   2383: 'Carrier 37 Encoder Comm Fault', class No Acknowledgement, trigger "DB302_HMI_Faults_Carrier37_Faults_0" bit 14
   2384: 'Carrier 37 HMI Comm Fault', class No Acknowledgement, trigger "DB302_HMI_Faults_Carrier37_Faults_0" bit 15
   2385: 'Carrier 37 Crash Detection Fault', class No Acknowledgement, trigger "DB302_HMI_Faults_Carrier37_Faults_1" bit 0
   2386: 'Carrier 37 Carrier Number Invalid', class No Acknowledgement, trigger "DB302_HMI_Faults_Carrier37_Faults_1" bit 1
   2387: 'Carrier 37 Drive: PROFINET configuration error', class No Acknowledgement, trigger "DB302_HMI_Faults_Carrier37_Faults_1" bit 2
   2388: 'Carrier 37 Drive: Error internal communications', class No Acknowledgement, trigger "DB302_HMI_Faults_Carrier37_Faults_1" bit 3
   2389: 'Carrier 37 Drive: Motor overtemperature', class No Acknowledgement, trigger "DB302_HMI_Faults_Carrier37_Faults_1" bit 4
   2390: 'Carrier 37 Drive: Motor overcurrent', class No Acknowledgement, trigger "DB302_HMI_Faults_Carrier37_Faults_1" bit 5
   2391: 'Carrier 37 Drive: Infeed or power unit not ready', class No Acknowledgement, trigger "DB302_HMI_Faults_Carrier37_Faults_1" bit 6
   2392: 'Carrier 37 Drive: Short-circuit/ground fault detected', class No Acknowledgement, trigger "DB302_HMI_Faults_Carrier37_Faults_1" bit 7
   2393: 'Carrier 37 Drive: PROFINET Setpoint timeout', class No Acknowledgement, trigger "DB302_HMI_Faults_Carrier37_Faults_1" bit 8
   2394: 'Carrier 37 Power unit: Overcurrent', class No Acknowledgement, trigger "DB302_HMI_Faults_Carrier37_Faults_1" bit 9
   2395: 'Carrier 37 Power unit: DC link voltage overvoltage', class No Acknowledgement, trigger "DB302_HMI_Faults_Carrier37_Faults_1" bit 10
   2396: 'Carrier 37 Power unit: DC link voltage undervoltage', class No Acknowledgement, trigger "DB302_HMI_Faults_Carrier37_Faults_1" bit 11
   2397: 'Carrier 37 Power unit: Line phase failure in main circuit', class No Acknowledgement, trigger "DB302_HMI_Faults_Carrier37_Faults_1" bit 12
   2398: 'Carrier 37 Power unit: Phase failure motor cable', class No Acknowledgement, trigger "DB302_HMI_Faults_Carrier37_Faults_1" bit 13
   2399: 'Carrier 37 Power unit: Ground fault', class No Acknowledgement, trigger "DB302_HMI_Faults_Carrier37_Faults_1" bit 14
   2400: 'Spare_Fault_2400', class No Acknowledgement, trigger "DB302_HMI_Faults_Carrier37_Faults_1" bit 15
   2401: 'Carrier 37 Motion Off Fault', class No Acknowledgement, trigger "DB302_HMI_Faults_Carrier37_Faults_2" bit 0
   2402: 'Carrier 37 Motion On Fault', class No Acknowledgement, trigger "DB302_HMI_Faults_Carrier37_Faults_2" bit 1
   2403: 'Carrier 37 Spacing Fault', class No Acknowledgement, trigger "DB302_HMI_Faults_Carrier37_Faults_2" bit 2
   2404: 'Carrier 37 Duplicate Carrier Number Fault', class No Acknowledgement, trigger "DB302_HMI_Faults_Carrier37_Faults_2" bit 3
   2405: 'Spare_Fault_2405', class No Acknowledgement, trigger "DB302_HMI_Faults_Carrier37_Faults_2" bit 4
   2406: 'Spare_Fault_2406', class No Acknowledgement, trigger "DB302_HMI_Faults_Carrier37_Faults_2" bit 5
   2407: 'Spare_Fault_2407', class No Acknowledgement, trigger "DB302_HMI_Faults_Carrier37_Faults_2" bit 6
   2408: 'Spare_Fault_2408', class No Acknowledgement, trigger "DB302_HMI_Faults_Carrier37_Faults_2" bit 7
   2409: 'Spare_Fault_2409', class No Acknowledgement, trigger "DB302_HMI_Faults_Carrier37_Faults_2" bit 8
   2410: 'Spare_Fault_2410', class No Acknowledgement, trigger "DB302_HMI_Faults_Carrier37_Faults_2" bit 9
   2411: 'Spare_Fault_2411', class No Acknowledgement, trigger "DB302_HMI_Faults_Carrier37_Faults_2" bit 10
   2412: 'Spare_Fault_2412', class No Acknowledgement, trigger "DB302_HMI_Faults_Carrier37_Faults_2" bit 11
   2413: 'Spare_Fault_2413', class No Acknowledgement, trigger "DB302_HMI_Faults_Carrier37_Faults_2" bit 12
   2414: 'Spare_Fault_2414', class No Acknowledgement, trigger "DB302_HMI_Faults_Carrier37_Faults_2" bit 13
   2415: 'Spare_Fault_2415', class No Acknowledgement, trigger "DB302_HMI_Faults_Carrier37_Faults_2" bit 14
   2416: 'Spare_Fault_2416', class No Acknowledgement, trigger "DB302_HMI_Faults_Carrier37_Faults_2" bit 15
   2417: 'Spare_Fault_2417', class No Acknowledgement, trigger "DB302_HMI_Faults_Carrier37_Faults_3" bit 0
   2418: 'Spare_Fault_2418', class No Acknowledgement, trigger "DB302_HMI_Faults_Carrier37_Faults_3" bit 1
   2419: 'Spare_Fault_2419', class No Acknowledgement, trigger "DB302_HMI_Faults_Carrier37_Faults_3" bit 2
   2420: 'Spare_Fault_2420', class No Acknowledgement, trigger "DB302_HMI_Faults_Carrier37_Faults_3" bit 3
   2421: 'Spare_Fault_2421', class No Acknowledgement, trigger "DB302_HMI_Faults_Carrier37_Faults_3" bit 4
   2422: 'Spare_Fault_2422', class No Acknowledgement, trigger "DB302_HMI_Faults_Carrier37_Faults_3" bit 5
   2423: 'Spare_Fault_2423', class No Acknowledgement, trigger "DB302_HMI_Faults_Carrier37_Faults_3" bit 6
   2424: 'Spare_Fault_2424', class No Acknowledgement, trigger "DB302_HMI_Faults_Carrier37_Faults_3" bit 7
   2425: 'Spare_Fault_2425', class No Acknowledgement, trigger "DB302_HMI_Faults_Carrier37_Faults_3" bit 8
   2426: 'Spare_Fault_2426', class No Acknowledgement, trigger "DB302_HMI_Faults_Carrier37_Faults_3" bit 9
   2427: 'Spare_Fault_2427', class No Acknowledgement, trigger "DB302_HMI_Faults_Carrier37_Faults_3" bit 10
   2428: 'Spare_Fault_2428', class No Acknowledgement, trigger "DB302_HMI_Faults_Carrier37_Faults_3" bit 11
   2429: 'Spare_Fault_2429', class No Acknowledgement, trigger "DB302_HMI_Faults_Carrier37_Faults_3" bit 12
   2430: 'Spare_Fault_2430', class No Acknowledgement, trigger "DB302_HMI_Faults_Carrier37_Faults_3" bit 13
   2431: 'Spare_Fault_2431', class No Acknowledgement, trigger "DB302_HMI_Faults_Carrier37_Faults_3" bit 14
   2432: 'Spare_Fault_2432', class No Acknowledgement, trigger "DB302_HMI_Faults_Carrier37_Faults_3" bit 15
   2433: 'Carrier 38 Disconnect Open Power Fault DI11.0', class No Acknowledgement, trigger "DB302_HMI_Faults_Carrier38_Faults_0" bit 0
   2434: 'Carrier 38 Drive Profinet Comm Fault', class No Acknowledgement, trigger "DB302_HMI_Faults_Carrier38_Faults_0" bit 1
   2435: 'Carrier 38 Production Stop Not Reset', class No Acknowledgement, trigger "DB302_HMI_Faults_Carrier38_Faults_0" bit 2
   2436: 'Carrier 38 CB02122 Tripped', class No Acknowledgement, trigger "DB302_HMI_Faults_Carrier38_Faults_0" bit 3
   2437: 'Carrier 38 CB02123 Tripped', class No Acknowledgement, trigger "DB302_HMI_Faults_Carrier38_Faults_0" bit 4
   2438: 'Carrier 38 AUX1 CB Tripped', class No Acknowledgement, trigger "DB302_HMI_Faults_Carrier38_Faults_0" bit 5
   2439: 'Carrier 38 AUX2 CB Tripped', class No Acknowledgement, trigger "DB302_HMI_Faults_Carrier38_Faults_0" bit 6
   2440: 'Carrier 38 PLC Not Communicating', class No Acknowledgement, trigger "DB302_HMI_Faults_Carrier38_Faults_0" bit 7
   2441: 'Carrier 38 Safe Input Card Fault', class No Acknowledgement, trigger "DB302_HMI_Faults_Carrier38_Faults_0" bit 8
   2442: 'Carrier 38 Safe Output Card Fault', class No Acknowledgement, trigger "DB302_HMI_Faults_Carrier38_Faults_0" bit 9
   2443: 'Carrier 38 Standard Input Card Fault', class No Acknowledgement, trigger "DB302_HMI_Faults_Carrier38_Faults_0" bit 10
   2444: 'Carrier 38 Standard Output Card Fault', class No Acknowledgement, trigger "DB302_HMI_Faults_Carrier38_Faults_0" bit 11
   2445: 'Carrier 38 Encoder Position Fault', class No Acknowledgement, trigger "DB302_HMI_Faults_Carrier38_Faults_0" bit 12
   2446: 'Carrier 38 Encoder Internal Error', class No Acknowledgement, trigger "DB302_HMI_Faults_Carrier38_Faults_0" bit 13
   2447: 'Carrier 38 Encoder Comm Fault', class No Acknowledgement, trigger "DB302_HMI_Faults_Carrier38_Faults_0" bit 14
   2448: 'Carrier 38 HMI Comm Fault', class No Acknowledgement, trigger "DB302_HMI_Faults_Carrier38_Faults_0" bit 15
   2449: 'Carrier 38 Crash Detection Fault', class No Acknowledgement, trigger "DB302_HMI_Faults_Carrier38_Faults_1" bit 0
   2450: 'Carrier 38 Carrier Number Invalid', class No Acknowledgement, trigger "DB302_HMI_Faults_Carrier38_Faults_1" bit 1
   2451: 'Carrier 38 Drive: PROFINET configuration error', class No Acknowledgement, trigger "DB302_HMI_Faults_Carrier38_Faults_1" bit 2
   2452: 'Carrier 38 Drive: Error internal communications', class No Acknowledgement, trigger "DB302_HMI_Faults_Carrier38_Faults_1" bit 3
   2453: 'Carrier 38 Drive: Motor overtemperature', class No Acknowledgement, trigger "DB302_HMI_Faults_Carrier38_Faults_1" bit 4
   2454: 'Carrier 38 Drive: Motor overcurrent', class No Acknowledgement, trigger "DB302_HMI_Faults_Carrier38_Faults_1" bit 5
   2455: 'Carrier 38 Drive: Infeed or power unit not ready', class No Acknowledgement, trigger "DB302_HMI_Faults_Carrier38_Faults_1" bit 6
   2456: 'Carrier 38 Drive: Short-circuit/ground fault detected', class No Acknowledgement, trigger "DB302_HMI_Faults_Carrier38_Faults_1" bit 7
   2457: 'Carrier 38 Drive: PROFINET Setpoint timeout', class No Acknowledgement, trigger "DB302_HMI_Faults_Carrier38_Faults_1" bit 8
   2458: 'Carrier 38 Power unit: Overcurrent', class No Acknowledgement, trigger "DB302_HMI_Faults_Carrier38_Faults_1" bit 9
   2459: 'Carrier 38 Power unit: DC link voltage overvoltage', class No Acknowledgement, trigger "DB302_HMI_Faults_Carrier38_Faults_1" bit 10
   2460: 'Carrier 38 Power unit: DC link voltage undervoltage', class No Acknowledgement, trigger "DB302_HMI_Faults_Carrier38_Faults_1" bit 11
   2461: 'Carrier 38 Power unit: Line phase failure in main circuit', class No Acknowledgement, trigger "DB302_HMI_Faults_Carrier38_Faults_1" bit 12
   2462: 'Carrier 38 Power unit: Phase failure motor cable', class No Acknowledgement, trigger "DB302_HMI_Faults_Carrier38_Faults_1" bit 13
   2463: 'Carrier 38 Power unit: Ground fault', class No Acknowledgement, trigger "DB302_HMI_Faults_Carrier38_Faults_1" bit 14
   2464: 'Spare_Fault_2464', class No Acknowledgement, trigger "DB302_HMI_Faults_Carrier38_Faults_1" bit 15
   2465: 'Carrier 38 Motion Off Fault', class No Acknowledgement, trigger "DB302_HMI_Faults_Carrier38_Faults_2" bit 0
   2466: 'Carrier 38 Motion On Fault', class No Acknowledgement, trigger "DB302_HMI_Faults_Carrier38_Faults_2" bit 1
   2467: 'Carrier 38 Spacing Fault', class No Acknowledgement, trigger "DB302_HMI_Faults_Carrier38_Faults_2" bit 2
   2468: 'Carrier 38 Duplicate Carrier Number Fault', class No Acknowledgement, trigger "DB302_HMI_Faults_Carrier38_Faults_2" bit 3
   2469: 'Spare_Fault_2469', class No Acknowledgement, trigger "DB302_HMI_Faults_Carrier38_Faults_2" bit 4
   2470: 'Spare_Fault_2470', class No Acknowledgement, trigger "DB302_HMI_Faults_Carrier38_Faults_2" bit 5
   2471: 'Spare_Fault_2471', class No Acknowledgement, trigger "DB302_HMI_Faults_Carrier38_Faults_2" bit 6
   2472: 'Spare_Fault_2472', class No Acknowledgement, trigger "DB302_HMI_Faults_Carrier38_Faults_2" bit 7
   2473: 'Spare_Fault_2473', class No Acknowledgement, trigger "DB302_HMI_Faults_Carrier38_Faults_2" bit 8
   2474: 'Spare_Fault_2474', class No Acknowledgement, trigger "DB302_HMI_Faults_Carrier38_Faults_2" bit 9
   2475: 'Spare_Fault_2475', class No Acknowledgement, trigger "DB302_HMI_Faults_Carrier38_Faults_2" bit 10
   2476: 'Spare_Fault_2476', class No Acknowledgement, trigger "DB302_HMI_Faults_Carrier38_Faults_2" bit 11
   2477: 'Spare_Fault_2477', class No Acknowledgement, trigger "DB302_HMI_Faults_Carrier38_Faults_2" bit 12
   2478: 'Spare_Fault_2478', class No Acknowledgement, trigger "DB302_HMI_Faults_Carrier38_Faults_2" bit 13
   2479: 'Spare_Fault_2479', class No Acknowledgement, trigger "DB302_HMI_Faults_Carrier38_Faults_2" bit 14
   2480: 'Spare_Fault_2480', class No Acknowledgement, trigger "DB302_HMI_Faults_Carrier38_Faults_2" bit 15
   2481: 'Spare_Fault_2481', class No Acknowledgement, trigger "DB302_HMI_Faults_Carrier38_Faults_3" bit 0
   2482: 'Spare_Fault_2482', class No Acknowledgement, trigger "DB302_HMI_Faults_Carrier38_Faults_3" bit 1
   2483: 'Spare_Fault_2483', class No Acknowledgement, trigger "DB302_HMI_Faults_Carrier38_Faults_3" bit 2
   2484: 'Spare_Fault_2484', class No Acknowledgement, trigger "DB302_HMI_Faults_Carrier38_Faults_3" bit 3
   2485: 'Spare_Fault_2485', class No Acknowledgement, trigger "DB302_HMI_Faults_Carrier38_Faults_3" bit 4
   2486: 'Spare_Fault_2486', class No Acknowledgement, trigger "DB302_HMI_Faults_Carrier38_Faults_3" bit 5
   2487: 'Spare_Fault_2487', class No Acknowledgement, trigger "DB302_HMI_Faults_Carrier38_Faults_3" bit 6
   2488: 'Spare_Fault_2488', class No Acknowledgement, trigger "DB302_HMI_Faults_Carrier38_Faults_3" bit 7
   2489: 'Spare_Fault_2489', class No Acknowledgement, trigger "DB302_HMI_Faults_Carrier38_Faults_3" bit 8
   2490: 'Spare_Fault_2490', class No Acknowledgement, trigger "DB302_HMI_Faults_Carrier38_Faults_3" bit 9
   2491: 'Spare_Fault_2491', class No Acknowledgement, trigger "DB302_HMI_Faults_Carrier38_Faults_3" bit 10
   2492: 'Spare_Fault_2492', class No Acknowledgement, trigger "DB302_HMI_Faults_Carrier38_Faults_3" bit 11
   2493: 'Spare_Fault_2493', class No Acknowledgement, trigger "DB302_HMI_Faults_Carrier38_Faults_3" bit 12
   2494: 'Spare_Fault_2494', class No Acknowledgement, trigger "DB302_HMI_Faults_Carrier38_Faults_3" bit 13
   2495: 'Spare_Fault_2495', class No Acknowledgement, trigger "DB302_HMI_Faults_Carrier38_Faults_3" bit 14
   2496: 'Spare_Fault_2496', class No Acknowledgement, trigger "DB302_HMI_Faults_Carrier38_Faults_3" bit 15
   2497: 'Carrier 39 Disconnect Open Power Fault DI11.0', class No Acknowledgement, trigger "DB302_HMI_Faults_Carrier39_Faults_0" bit 0
   2498: 'Carrier 39 Drive Profinet Comm Fault', class No Acknowledgement, trigger "DB302_HMI_Faults_Carrier39_Faults_0" bit 1
   2499: 'Carrier 39 Production Stop Not Reset', class No Acknowledgement, trigger "DB302_HMI_Faults_Carrier39_Faults_0" bit 2
   2500: 'Carrier 39 CB02122 Tripped', class No Acknowledgement, trigger "DB302_HMI_Faults_Carrier39_Faults_0" bit 3
   2501: 'Carrier 39 CB02123 Tripped', class No Acknowledgement, trigger "DB302_HMI_Faults_Carrier39_Faults_0" bit 4
   2502: 'Carrier 39 AUX1 CB Tripped', class No Acknowledgement, trigger "DB302_HMI_Faults_Carrier39_Faults_0" bit 5
   2503: 'Carrier 39 AUX2 CB Tripped', class No Acknowledgement, trigger "DB302_HMI_Faults_Carrier39_Faults_0" bit 6
   2504: 'Carrier 39 PLC Not Communicating', class No Acknowledgement, trigger "DB302_HMI_Faults_Carrier39_Faults_0" bit 7
   2505: 'Carrier 39 Safe Input Card Fault', class No Acknowledgement, trigger "DB302_HMI_Faults_Carrier39_Faults_0" bit 8
   2506: 'Carrier 39 Safe Output Card Fault', class No Acknowledgement, trigger "DB302_HMI_Faults_Carrier39_Faults_0" bit 9
   2507: 'Carrier 39 Standard Input Card Fault', class No Acknowledgement, trigger "DB302_HMI_Faults_Carrier39_Faults_0" bit 10
   2508: 'Carrier 39 Standard Output Card Fault', class No Acknowledgement, trigger "DB302_HMI_Faults_Carrier39_Faults_0" bit 11
   2509: 'Carrier 39 Encoder Position Fault', class No Acknowledgement, trigger "DB302_HMI_Faults_Carrier39_Faults_0" bit 12
   2510: 'Carrier 39 Encoder Internal Error', class No Acknowledgement, trigger "DB302_HMI_Faults_Carrier39_Faults_0" bit 13
   2511: 'Carrier 39 Encoder Comm Fault', class No Acknowledgement, trigger "DB302_HMI_Faults_Carrier39_Faults_0" bit 14
   2512: 'Carrier 39 HMI Comm Fault', class No Acknowledgement, trigger "DB302_HMI_Faults_Carrier39_Faults_0" bit 15
   2513: 'Carrier 39 Crash Detection Fault', class No Acknowledgement, trigger "DB302_HMI_Faults_Carrier39_Faults_1" bit 0
   2514: 'Carrier 39 Carrier Number Invalid', class No Acknowledgement, trigger "DB302_HMI_Faults_Carrier39_Faults_1" bit 1
   2515: 'Carrier 39 Drive: PROFINET configuration error', class No Acknowledgement, trigger "DB302_HMI_Faults_Carrier39_Faults_1" bit 2
   2516: 'Carrier 39 Drive: Error internal communications', class No Acknowledgement, trigger "DB302_HMI_Faults_Carrier39_Faults_1" bit 3
   2517: 'Carrier 39 Drive: Motor overtemperature', class No Acknowledgement, trigger "DB302_HMI_Faults_Carrier39_Faults_1" bit 4
   2518: 'Carrier 39 Drive: Motor overcurrent', class No Acknowledgement, trigger "DB302_HMI_Faults_Carrier39_Faults_1" bit 5
   2519: 'Carrier 39 Drive: Infeed or power unit not ready', class No Acknowledgement, trigger "DB302_HMI_Faults_Carrier39_Faults_1" bit 6
   2520: 'Carrier 39 Drive: Short-circuit/ground fault detected', class No Acknowledgement, trigger "DB302_HMI_Faults_Carrier39_Faults_1" bit 7
   2521: 'Carrier 39 Drive: PROFINET Setpoint timeout', class No Acknowledgement, trigger "DB302_HMI_Faults_Carrier39_Faults_1" bit 8
   2522: 'Carrier 39 Power unit: Overcurrent', class No Acknowledgement, trigger "DB302_HMI_Faults_Carrier39_Faults_1" bit 9
   2523: 'Carrier 39 Power unit: DC link voltage overvoltage', class No Acknowledgement, trigger "DB302_HMI_Faults_Carrier39_Faults_1" bit 10
   2524: 'Carrier 39 Power unit: DC link voltage undervoltage', class No Acknowledgement, trigger "DB302_HMI_Faults_Carrier39_Faults_1" bit 11
   2525: 'Carrier 39 Power unit: Line phase failure in main circuit', class No Acknowledgement, trigger "DB302_HMI_Faults_Carrier39_Faults_1" bit 12
   2526: 'Carrier 39 Power unit: Phase failure motor cable', class No Acknowledgement, trigger "DB302_HMI_Faults_Carrier39_Faults_1" bit 13
   2527: 'Carrier 39 Power unit: Ground fault', class No Acknowledgement, trigger "DB302_HMI_Faults_Carrier39_Faults_1" bit 14
   2528: 'Spare_Fault_2528', class No Acknowledgement, trigger "DB302_HMI_Faults_Carrier39_Faults_1" bit 15
   2529: 'Carrier 39 Motion Off Fault', class No Acknowledgement, trigger "DB302_HMI_Faults_Carrier39_Faults_2" bit 0
   2530: 'Carrier 39 Motion On Fault', class No Acknowledgement, trigger "DB302_HMI_Faults_Carrier39_Faults_2" bit 1
   2531: 'Carrier 39 Spacing Fault', class No Acknowledgement, trigger "DB302_HMI_Faults_Carrier39_Faults_2" bit 2
   2532: 'Carrier 39 Duplicate Carrier Number Fault', class No Acknowledgement, trigger "DB302_HMI_Faults_Carrier39_Faults_2" bit 3
   2533: 'Spare_Fault_2533', class No Acknowledgement, trigger "DB302_HMI_Faults_Carrier39_Faults_2" bit 4
   2534: 'Spare_Fault_2534', class No Acknowledgement, trigger "DB302_HMI_Faults_Carrier39_Faults_2" bit 5
   2535: 'Spare_Fault_2535', class No Acknowledgement, trigger "DB302_HMI_Faults_Carrier39_Faults_2" bit 6
   2536: 'Spare_Fault_2536', class No Acknowledgement, trigger "DB302_HMI_Faults_Carrier39_Faults_2" bit 7
   2537: 'Spare_Fault_2537', class No Acknowledgement, trigger "DB302_HMI_Faults_Carrier39_Faults_2" bit 8
   2538: 'Spare_Fault_2538', class No Acknowledgement, trigger "DB302_HMI_Faults_Carrier39_Faults_2" bit 9
   2539: 'Spare_Fault_2539', class No Acknowledgement, trigger "DB302_HMI_Faults_Carrier39_Faults_2" bit 10
   2540: 'Spare_Fault_2540', class No Acknowledgement, trigger "DB302_HMI_Faults_Carrier39_Faults_2" bit 11
   2541: 'Spare_Fault_2541', class No Acknowledgement, trigger "DB302_HMI_Faults_Carrier39_Faults_2" bit 12
   2542: 'Spare_Fault_2542', class No Acknowledgement, trigger "DB302_HMI_Faults_Carrier39_Faults_2" bit 13
   2543: 'Spare_Fault_2543', class No Acknowledgement, trigger "DB302_HMI_Faults_Carrier39_Faults_2" bit 14
   2544: 'Spare_Fault_2544', class No Acknowledgement, trigger "DB302_HMI_Faults_Carrier39_Faults_2" bit 15
   2545: 'Spare_Fault_2545', class No Acknowledgement, trigger "DB302_HMI_Faults_Carrier39_Faults_3" bit 0
   2546: 'Spare_Fault_2546', class No Acknowledgement, trigger "DB302_HMI_Faults_Carrier39_Faults_3" bit 1
   2547: 'Spare_Fault_2547', class No Acknowledgement, trigger "DB302_HMI_Faults_Carrier39_Faults_3" bit 2
   2548: 'Spare_Fault_2548', class No Acknowledgement, trigger "DB302_HMI_Faults_Carrier39_Faults_3" bit 3
   2549: 'Spare_Fault_2549', class No Acknowledgement, trigger "DB302_HMI_Faults_Carrier39_Faults_3" bit 4
   2550: 'Spare_Fault_2550', class No Acknowledgement, trigger "DB302_HMI_Faults_Carrier39_Faults_3" bit 5
   2551: 'Spare_Fault_2551', class No Acknowledgement, trigger "DB302_HMI_Faults_Carrier39_Faults_3" bit 6
   2552: 'Spare_Fault_2552', class No Acknowledgement, trigger "DB302_HMI_Faults_Carrier39_Faults_3" bit 7
   2553: 'Spare_Fault_2553', class No Acknowledgement, trigger "DB302_HMI_Faults_Carrier39_Faults_3" bit 8
   2554: 'Spare_Fault_2554', class No Acknowledgement, trigger "DB302_HMI_Faults_Carrier39_Faults_3" bit 9
   2555: 'Spare_Fault_2555', class No Acknowledgement, trigger "DB302_HMI_Faults_Carrier39_Faults_3" bit 10
   2556: 'Spare_Fault_2556', class No Acknowledgement, trigger "DB302_HMI_Faults_Carrier39_Faults_3" bit 11
   2557: 'Spare_Fault_2557', class No Acknowledgement, trigger "DB302_HMI_Faults_Carrier39_Faults_3" bit 12
   2558: 'Spare_Fault_2558', class No Acknowledgement, trigger "DB302_HMI_Faults_Carrier39_Faults_3" bit 13
   2559: 'Spare_Fault_2559', class No Acknowledgement, trigger "DB302_HMI_Faults_Carrier39_Faults_3" bit 14
   2560: 'Spare_Fault_2560', class No Acknowledgement, trigger "DB302_HMI_Faults_Carrier39_Faults_3" bit 15
   2561: 'Carrier 40 Disconnect Open Power Fault DI11.0', class No Acknowledgement, trigger "DB302_HMI_Faults_Carrier40_Faults_0" bit 0
   2562: 'Carrier 40 Drive Profinet Comm Fault', class No Acknowledgement, trigger "DB302_HMI_Faults_Carrier40_Faults_0" bit 1
   2563: 'Carrier 40 Production Stop Not Reset', class No Acknowledgement, trigger "DB302_HMI_Faults_Carrier40_Faults_0" bit 2
   2564: 'Carrier 40 CB02122 Tripped', class No Acknowledgement, trigger "DB302_HMI_Faults_Carrier40_Faults_0" bit 3
   2565: 'Carrier 40 CB02123 Tripped', class No Acknowledgement, trigger "DB302_HMI_Faults_Carrier40_Faults_0" bit 4
   2566: 'Carrier 40 AUX1 CB Tripped', class No Acknowledgement, trigger "DB302_HMI_Faults_Carrier40_Faults_0" bit 5
   2567: 'Carrier 40 AUX2 CB Tripped', class No Acknowledgement, trigger "DB302_HMI_Faults_Carrier40_Faults_0" bit 6
   2568: 'Carrier 40 PLC Not Communicating', class No Acknowledgement, trigger "DB302_HMI_Faults_Carrier40_Faults_0" bit 7
   2569: 'Carrier 40 Safe Input Card Fault', class No Acknowledgement, trigger "DB302_HMI_Faults_Carrier40_Faults_0" bit 8
   2570: 'Carrier 40 Safe Output Card Fault', class No Acknowledgement, trigger "DB302_HMI_Faults_Carrier40_Faults_0" bit 9
   2571: 'Carrier 40 Standard Input Card Fault', class No Acknowledgement, trigger "DB302_HMI_Faults_Carrier40_Faults_0" bit 10
   2572: 'Carrier 40 Standard Output Card Fault', class No Acknowledgement, trigger "DB302_HMI_Faults_Carrier40_Faults_0" bit 11
   2573: 'Carrier 40 Encoder Position Fault', class No Acknowledgement, trigger "DB302_HMI_Faults_Carrier40_Faults_0" bit 12
   2574: 'Carrier 40 Encoder Internal Error', class No Acknowledgement, trigger "DB302_HMI_Faults_Carrier40_Faults_0" bit 13
   2575: 'Carrier 40 Encoder Comm Fault', class No Acknowledgement, trigger "DB302_HMI_Faults_Carrier40_Faults_0" bit 14
   2576: 'Carrier 40 HMI Comm Fault', class No Acknowledgement, trigger "DB302_HMI_Faults_Carrier40_Faults_0" bit 15
   2577: 'Carrier 40 Crash Detection Fault', class No Acknowledgement, trigger "DB302_HMI_Faults_Carrier40_Faults_1" bit 0
   2578: 'Carrier 40 Carrier Number Invalid', class No Acknowledgement, trigger "DB302_HMI_Faults_Carrier40_Faults_1" bit 1
   2579: 'Carrier 40 Drive: PROFINET configuration error', class No Acknowledgement, trigger "DB302_HMI_Faults_Carrier40_Faults_1" bit 2
   2580: 'Carrier 40 Drive: Error internal communications', class No Acknowledgement, trigger "DB302_HMI_Faults_Carrier40_Faults_1" bit 3
   2581: 'Carrier 40 Drive: Motor overtemperature', class No Acknowledgement, trigger "DB302_HMI_Faults_Carrier40_Faults_1" bit 4
   2582: 'Carrier 40 Drive: Motor overcurrent', class No Acknowledgement, trigger "DB302_HMI_Faults_Carrier40_Faults_1" bit 5
   2583: 'Carrier 40 Drive: Infeed or power unit not ready', class No Acknowledgement, trigger "DB302_HMI_Faults_Carrier40_Faults_1" bit 6
   2584: 'Carrier 40 Drive: Short-circuit/ground fault detected', class No Acknowledgement, trigger "DB302_HMI_Faults_Carrier40_Faults_1" bit 7
   2585: 'Carrier 40 Drive: PROFINET Setpoint timeout', class No Acknowledgement, trigger "DB302_HMI_Faults_Carrier40_Faults_1" bit 8
   2586: 'Carrier 40 Power unit: Overcurrent', class No Acknowledgement, trigger "DB302_HMI_Faults_Carrier40_Faults_1" bit 9
   2587: 'Carrier 40 Power unit: DC link voltage overvoltage', class No Acknowledgement, trigger "DB302_HMI_Faults_Carrier40_Faults_1" bit 10
   2588: 'Carrier 40 Power unit: DC link voltage undervoltage', class No Acknowledgement, trigger "DB302_HMI_Faults_Carrier40_Faults_1" bit 11
   2589: 'Carrier 40 Power unit: Line phase failure in main circuit', class No Acknowledgement, trigger "DB302_HMI_Faults_Carrier40_Faults_1" bit 12
   2590: 'Carrier 40 Power unit: Phase failure motor cable', class No Acknowledgement, trigger "DB302_HMI_Faults_Carrier40_Faults_1" bit 13
   2591: 'Carrier 40 Power unit: Ground fault', class No Acknowledgement, trigger "DB302_HMI_Faults_Carrier40_Faults_1" bit 14
   2592: 'Spare_Fault_2592', class No Acknowledgement, trigger "DB302_HMI_Faults_Carrier40_Faults_1" bit 15
   2593: 'Carrier 40 Motion Off Fault', class No Acknowledgement, trigger "DB302_HMI_Faults_Carrier40_Faults_2" bit 0
   2594: 'Carrier 40 Motion On Fault', class No Acknowledgement, trigger "DB302_HMI_Faults_Carrier40_Faults_2" bit 1
   2595: 'Carrier 40 Spacing Fault', class No Acknowledgement, trigger "DB302_HMI_Faults_Carrier40_Faults_2" bit 2
   2596: 'Carrier 40 Duplicate Carrier Number Fault', class No Acknowledgement, trigger "DB302_HMI_Faults_Carrier40_Faults_2" bit 3
   2597: 'Spare_Fault_2597', class No Acknowledgement, trigger "DB302_HMI_Faults_Carrier40_Faults_2" bit 4
   2598: 'Spare_Fault_2598', class No Acknowledgement, trigger "DB302_HMI_Faults_Carrier40_Faults_2" bit 5
   2599: 'Spare_Fault_2599', class No Acknowledgement, trigger "DB302_HMI_Faults_Carrier40_Faults_2" bit 6
   2600: 'Spare_Fault_2600', class No Acknowledgement, trigger "DB302_HMI_Faults_Carrier40_Faults_2" bit 7
   2601: 'Spare_Fault_2601', class No Acknowledgement, trigger "DB302_HMI_Faults_Carrier40_Faults_2" bit 8
   2602: 'Spare_Fault_2602', class No Acknowledgement, trigger "DB302_HMI_Faults_Carrier40_Faults_2" bit 9
   2603: 'Spare_Fault_2603', class No Acknowledgement, trigger "DB302_HMI_Faults_Carrier40_Faults_2" bit 10
   2604: 'Spare_Fault_2604', class No Acknowledgement, trigger "DB302_HMI_Faults_Carrier40_Faults_2" bit 11
   2605: 'Spare_Fault_2605', class No Acknowledgement, trigger "DB302_HMI_Faults_Carrier40_Faults_2" bit 12
   2606: 'Spare_Fault_2606', class No Acknowledgement, trigger "DB302_HMI_Faults_Carrier40_Faults_2" bit 13
   2607: 'Spare_Fault_2607', class No Acknowledgement, trigger "DB302_HMI_Faults_Carrier40_Faults_2" bit 14
   2608: 'Spare_Fault_2608', class No Acknowledgement, trigger "DB302_HMI_Faults_Carrier40_Faults_2" bit 15
   2609: 'Spare_Fault_2609', class No Acknowledgement, trigger "DB302_HMI_Faults_Carrier40_Faults_3" bit 0
   2610: 'Spare_Fault_2610', class No Acknowledgement, trigger "DB302_HMI_Faults_Carrier40_Faults_3" bit 1
   2611: 'Spare_Fault_2611', class No Acknowledgement, trigger "DB302_HMI_Faults_Carrier40_Faults_3" bit 2
   2612: 'Spare_Fault_2612', class No Acknowledgement, trigger "DB302_HMI_Faults_Carrier40_Faults_3" bit 3
   2613: 'Spare_Fault_2613', class No Acknowledgement, trigger "DB302_HMI_Faults_Carrier40_Faults_3" bit 4
   2614: 'Spare_Fault_2614', class No Acknowledgement, trigger "DB302_HMI_Faults_Carrier40_Faults_3" bit 5
   2615: 'Spare_Fault_2615', class No Acknowledgement, trigger "DB302_HMI_Faults_Carrier40_Faults_3" bit 6
   2616: 'Spare_Fault_2616', class No Acknowledgement, trigger "DB302_HMI_Faults_Carrier40_Faults_3" bit 7
   2617: 'Spare_Fault_2617', class No Acknowledgement, trigger "DB302_HMI_Faults_Carrier40_Faults_3" bit 8
   2618: 'Spare_Fault_2618', class No Acknowledgement, trigger "DB302_HMI_Faults_Carrier40_Faults_3" bit 9
   2619: 'Spare_Fault_2619', class No Acknowledgement, trigger "DB302_HMI_Faults_Carrier40_Faults_3" bit 10
   2620: 'Spare_Fault_2620', class No Acknowledgement, trigger "DB302_HMI_Faults_Carrier40_Faults_3" bit 11
   2621: 'Spare_Fault_2621', class No Acknowledgement, trigger "DB302_HMI_Faults_Carrier40_Faults_3" bit 12
   2622: 'Spare_Fault_2622', class No Acknowledgement, trigger "DB302_HMI_Faults_Carrier40_Faults_3" bit 13
   2623: 'Spare_Fault_2623', class No Acknowledgement, trigger "DB302_HMI_Faults_Carrier40_Faults_3" bit 14
   2624: 'Spare_Fault_2624', class No Acknowledgement, trigger "DB302_HMI_Faults_Carrier40_Faults_3" bit 15
   2625: 'Carrier 41 Disconnect Open Power Fault DI11.0', class No Acknowledgement, trigger "DB302_HMI_Faults_Carrier41_Faults_0" bit 0
   2626: 'Carrier 41 Drive Profinet Comm Fault', class No Acknowledgement, trigger "DB302_HMI_Faults_Carrier41_Faults_0" bit 1
   2627: 'Carrier 41 Production Stop Not Reset', class No Acknowledgement, trigger "DB302_HMI_Faults_Carrier41_Faults_0" bit 2
   2628: 'Carrier 41 CB02122 Tripped', class No Acknowledgement, trigger "DB302_HMI_Faults_Carrier41_Faults_0" bit 3
   2629: 'Carrier 41 CB02123 Tripped', class No Acknowledgement, trigger "DB302_HMI_Faults_Carrier41_Faults_0" bit 4
   2630: 'Carrier 41 AUX1 CB Tripped', class No Acknowledgement, trigger "DB302_HMI_Faults_Carrier41_Faults_0" bit 5
   2631: 'Carrier 41 AUX2 CB Tripped', class No Acknowledgement, trigger "DB302_HMI_Faults_Carrier41_Faults_0" bit 6
   2632: 'Carrier 41 PLC Not Communicating', class No Acknowledgement, trigger "DB302_HMI_Faults_Carrier41_Faults_0" bit 7
   2633: 'Carrier 41 Safe Input Card Fault', class No Acknowledgement, trigger "DB302_HMI_Faults_Carrier41_Faults_0" bit 8
   2634: 'Carrier 41 Safe Output Card Fault', class No Acknowledgement, trigger "DB302_HMI_Faults_Carrier41_Faults_0" bit 9
   2635: 'Carrier 41 Standard Input Card Fault', class No Acknowledgement, trigger "DB302_HMI_Faults_Carrier41_Faults_0" bit 10
   2636: 'Carrier 41 Standard Output Card Fault', class No Acknowledgement, trigger "DB302_HMI_Faults_Carrier41_Faults_0" bit 11
   2637: 'Carrier 41 Encoder Position Fault', class No Acknowledgement, trigger "DB302_HMI_Faults_Carrier41_Faults_0" bit 12
   2638: 'Carrier 41 Encoder Internal Error', class No Acknowledgement, trigger "DB302_HMI_Faults_Carrier41_Faults_0" bit 13
   2639: 'Carrier 41 Encoder Comm Fault', class No Acknowledgement, trigger "DB302_HMI_Faults_Carrier41_Faults_0" bit 14
   2640: 'Carrier 41 HMI Comm Fault', class No Acknowledgement, trigger "DB302_HMI_Faults_Carrier41_Faults_0" bit 15
   2641: 'Carrier 41 Crash Detection Fault', class No Acknowledgement, trigger "DB302_HMI_Faults_Carrier41_Faults_1" bit 0
   2642: 'Carrier 41 Carrier Number Invalid', class No Acknowledgement, trigger "DB302_HMI_Faults_Carrier41_Faults_1" bit 1
   2643: 'Carrier 41 Drive: PROFINET configuration error', class No Acknowledgement, trigger "DB302_HMI_Faults_Carrier41_Faults_1" bit 2
   2644: 'Carrier 41 Drive: Error internal communications', class No Acknowledgement, trigger "DB302_HMI_Faults_Carrier41_Faults_1" bit 3
   2645: 'Carrier 41 Drive: Motor overtemperature', class No Acknowledgement, trigger "DB302_HMI_Faults_Carrier41_Faults_1" bit 4
   2646: 'Carrier 41 Drive: Motor overcurrent', class No Acknowledgement, trigger "DB302_HMI_Faults_Carrier41_Faults_1" bit 5
   2647: 'Carrier 41 Drive: Infeed or power unit not ready', class No Acknowledgement, trigger "DB302_HMI_Faults_Carrier41_Faults_1" bit 6
   2648: 'Carrier 41 Drive: Short-circuit/ground fault detected', class No Acknowledgement, trigger "DB302_HMI_Faults_Carrier41_Faults_1" bit 7
   2649: 'Carrier 41 Drive: PROFINET Setpoint timeout', class No Acknowledgement, trigger "DB302_HMI_Faults_Carrier41_Faults_1" bit 8
   2650: 'Carrier 41 Power unit: Overcurrent', class No Acknowledgement, trigger "DB302_HMI_Faults_Carrier41_Faults_1" bit 9
   2651: 'Carrier 41 Power unit: DC link voltage overvoltage', class No Acknowledgement, trigger "DB302_HMI_Faults_Carrier41_Faults_1" bit 10
   2652: 'Carrier 41 Power unit: DC link voltage undervoltage', class No Acknowledgement, trigger "DB302_HMI_Faults_Carrier41_Faults_1" bit 11
   2653: 'Carrier 41 Power unit: Line phase failure in main circuit', class No Acknowledgement, trigger "DB302_HMI_Faults_Carrier41_Faults_1" bit 12
   2654: 'Carrier 41 Power unit: Phase failure motor cable', class No Acknowledgement, trigger "DB302_HMI_Faults_Carrier41_Faults_1" bit 13
   2655: 'Carrier 41 Power unit: Ground fault', class No Acknowledgement, trigger "DB302_HMI_Faults_Carrier41_Faults_1" bit 14
   2656: 'Spare_Fault_2656', class No Acknowledgement, trigger "DB302_HMI_Faults_Carrier41_Faults_1" bit 15
   2657: 'Carrier 41 Motion Off Fault', class No Acknowledgement, trigger "DB302_HMI_Faults_Carrier41_Faults_2" bit 0
   2658: 'Carrier 41 Motion On Fault', class No Acknowledgement, trigger "DB302_HMI_Faults_Carrier41_Faults_2" bit 1
   2659: 'Carrier 41 Spacing Fault', class No Acknowledgement, trigger "DB302_HMI_Faults_Carrier41_Faults_2" bit 2
   2660: 'Carrier 41 Duplicate Carrier Number Fault', class No Acknowledgement, trigger "DB302_HMI_Faults_Carrier41_Faults_2" bit 3
   2661: 'Spare_Fault_2661', class No Acknowledgement, trigger "DB302_HMI_Faults_Carrier41_Faults_2" bit 4
   2662: 'Spare_Fault_2662', class No Acknowledgement, trigger "DB302_HMI_Faults_Carrier41_Faults_2" bit 5
   2663: 'Spare_Fault_2663', class No Acknowledgement, trigger "DB302_HMI_Faults_Carrier41_Faults_2" bit 6
   2664: 'Spare_Fault_2664', class No Acknowledgement, trigger "DB302_HMI_Faults_Carrier41_Faults_2" bit 7
   2665: 'Spare_Fault_2665', class No Acknowledgement, trigger "DB302_HMI_Faults_Carrier41_Faults_2" bit 8
   2666: 'Spare_Fault_2666', class No Acknowledgement, trigger "DB302_HMI_Faults_Carrier41_Faults_2" bit 9
   2667: 'Spare_Fault_2667', class No Acknowledgement, trigger "DB302_HMI_Faults_Carrier41_Faults_2" bit 10
   2668: 'Spare_Fault_2668', class No Acknowledgement, trigger "DB302_HMI_Faults_Carrier41_Faults_2" bit 11
   2669: 'Spare_Fault_2669', class No Acknowledgement, trigger "DB302_HMI_Faults_Carrier41_Faults_2" bit 12
   2670: 'Spare_Fault_2670', class No Acknowledgement, trigger "DB302_HMI_Faults_Carrier41_Faults_2" bit 13
   2671: 'Spare_Fault_2671', class No Acknowledgement, trigger "DB302_HMI_Faults_Carrier41_Faults_2" bit 14
   2672: 'Spare_Fault_2672', class No Acknowledgement, trigger "DB302_HMI_Faults_Carrier41_Faults_2" bit 15
   2673: 'Spare_Fault_2673', class No Acknowledgement, trigger "DB302_HMI_Faults_Carrier41_Faults_3" bit 0
   2674: 'Spare_Fault_2674', class No Acknowledgement, trigger "DB302_HMI_Faults_Carrier41_Faults_3" bit 1
   2675: 'Spare_Fault_2675', class No Acknowledgement, trigger "DB302_HMI_Faults_Carrier41_Faults_3" bit 2
   2676: 'Spare_Fault_2676', class No Acknowledgement, trigger "DB302_HMI_Faults_Carrier41_Faults_3" bit 3
   2677: 'Spare_Fault_2677', class No Acknowledgement, trigger "DB302_HMI_Faults_Carrier41_Faults_3" bit 4
   2678: 'Spare_Fault_2678', class No Acknowledgement, trigger "DB302_HMI_Faults_Carrier41_Faults_3" bit 5
   2679: 'Spare_Fault_2679', class No Acknowledgement, trigger "DB302_HMI_Faults_Carrier41_Faults_3" bit 6
   2680: 'Spare_Fault_2680', class No Acknowledgement, trigger "DB302_HMI_Faults_Carrier41_Faults_3" bit 7
   2681: 'Spare_Fault_2681', class No Acknowledgement, trigger "DB302_HMI_Faults_Carrier41_Faults_3" bit 8
   2682: 'Spare_Fault_2682', class No Acknowledgement, trigger "DB302_HMI_Faults_Carrier41_Faults_3" bit 9
   2683: 'Spare_Fault_2683', class No Acknowledgement, trigger "DB302_HMI_Faults_Carrier41_Faults_3" bit 10
   2684: 'Spare_Fault_2684', class No Acknowledgement, trigger "DB302_HMI_Faults_Carrier41_Faults_3" bit 11
   2685: 'Spare_Fault_2685', class No Acknowledgement, trigger "DB302_HMI_Faults_Carrier41_Faults_3" bit 12
   2686: 'Spare_Fault_2686', class No Acknowledgement, trigger "DB302_HMI_Faults_Carrier41_Faults_3" bit 13
   2687: 'Spare_Fault_2687', class No Acknowledgement, trigger "DB302_HMI_Faults_Carrier41_Faults_3" bit 14
   2688: 'Spare_Fault_2688', class No Acknowledgement, trigger "DB302_HMI_Faults_Carrier41_Faults_3" bit 15
   2689: 'Carrier 42 Disconnect Open Power Fault DI11.0', class No Acknowledgement, trigger "DB302_HMI_Faults_Carrier42_Faults_0" bit 0
   2690: 'Carrier 42 Drive Profinet Comm Fault', class No Acknowledgement, trigger "DB302_HMI_Faults_Carrier42_Faults_0" bit 1
   2691: 'Carrier 42 Production Stop Not Reset', class No Acknowledgement, trigger "DB302_HMI_Faults_Carrier42_Faults_0" bit 2
   2692: 'Carrier 42 CB02122 Tripped', class No Acknowledgement, trigger "DB302_HMI_Faults_Carrier42_Faults_0" bit 3
   2693: 'Carrier 42 CB02123 Tripped', class No Acknowledgement, trigger "DB302_HMI_Faults_Carrier42_Faults_0" bit 4
   2694: 'Carrier 42 AUX1 CB Tripped', class No Acknowledgement, trigger "DB302_HMI_Faults_Carrier42_Faults_0" bit 5
   2695: 'Carrier 42 AUX2 CB Tripped', class No Acknowledgement, trigger "DB302_HMI_Faults_Carrier42_Faults_0" bit 6
   2696: 'Carrier 42 PLC Not Communicating', class No Acknowledgement, trigger "DB302_HMI_Faults_Carrier42_Faults_0" bit 7
   2697: 'Carrier 42 Safe Input Card Fault', class No Acknowledgement, trigger "DB302_HMI_Faults_Carrier42_Faults_0" bit 8
   2698: 'Carrier 42 Safe Output Card Fault', class No Acknowledgement, trigger "DB302_HMI_Faults_Carrier42_Faults_0" bit 9
   2699: 'Carrier 42 Standard Input Card Fault', class No Acknowledgement, trigger "DB302_HMI_Faults_Carrier42_Faults_0" bit 10
   2700: 'Carrier 42 Standard Output Card Fault', class No Acknowledgement, trigger "DB302_HMI_Faults_Carrier42_Faults_0" bit 11
   2701: 'Carrier 42 Encoder Position Fault', class No Acknowledgement, trigger "DB302_HMI_Faults_Carrier42_Faults_0" bit 12
   2702: 'Carrier 42 Encoder Internal Error', class No Acknowledgement, trigger "DB302_HMI_Faults_Carrier42_Faults_0" bit 13
   2703: 'Carrier 42 Encoder Comm Fault', class No Acknowledgement, trigger "DB302_HMI_Faults_Carrier42_Faults_0" bit 14
   2704: 'Carrier 42 HMI Comm Fault', class No Acknowledgement, trigger "DB302_HMI_Faults_Carrier42_Faults_0" bit 15
   2705: 'Carrier 42 Crash Detection Fault', class No Acknowledgement, trigger "DB302_HMI_Faults_Carrier42_Faults_1" bit 0
   2706: 'Carrier 42 Carrier Number Invalid', class No Acknowledgement, trigger "DB302_HMI_Faults_Carrier42_Faults_1" bit 1
   2707: 'Carrier 42 Drive: PROFINET configuration error', class No Acknowledgement, trigger "DB302_HMI_Faults_Carrier42_Faults_1" bit 2
   2708: 'Carrier 42 Drive: Error internal communications', class No Acknowledgement, trigger "DB302_HMI_Faults_Carrier42_Faults_1" bit 3
   2709: 'Carrier 42 Drive: Motor overtemperature', class No Acknowledgement, trigger "DB302_HMI_Faults_Carrier42_Faults_1" bit 4
   2710: 'Carrier 42 Drive: Motor overcurrent', class No Acknowledgement, trigger "DB302_HMI_Faults_Carrier42_Faults_1" bit 5
   2711: 'Carrier 42 Drive: Infeed or power unit not ready', class No Acknowledgement, trigger "DB302_HMI_Faults_Carrier42_Faults_1" bit 6
   2712: 'Carrier 42 Drive: Short-circuit/ground fault detected', class No Acknowledgement, trigger "DB302_HMI_Faults_Carrier42_Faults_1" bit 7
   2713: 'Carrier 42 Drive: PROFINET Setpoint timeout', class No Acknowledgement, trigger "DB302_HMI_Faults_Carrier42_Faults_1" bit 8
   2714: 'Carrier 42 Power unit: Overcurrent', class No Acknowledgement, trigger "DB302_HMI_Faults_Carrier42_Faults_1" bit 9
   2715: 'Carrier 42 Power unit: DC link voltage overvoltage', class No Acknowledgement, trigger "DB302_HMI_Faults_Carrier42_Faults_1" bit 10
   2716: 'Carrier 42 Power unit: DC link voltage undervoltage', class No Acknowledgement, trigger "DB302_HMI_Faults_Carrier42_Faults_1" bit 11
   2717: 'Carrier 42 Power unit: Line phase failure in main circuit', class No Acknowledgement, trigger "DB302_HMI_Faults_Carrier42_Faults_1" bit 12
   2718: 'Carrier 42 Power unit: Phase failure motor cable', class No Acknowledgement, trigger "DB302_HMI_Faults_Carrier42_Faults_1" bit 13
   2719: 'Carrier 42 Power unit: Ground fault', class No Acknowledgement, trigger "DB302_HMI_Faults_Carrier42_Faults_1" bit 14
   2720: 'Spare_Fault_2720', class No Acknowledgement, trigger "DB302_HMI_Faults_Carrier42_Faults_1" bit 15
   2721: 'Carrier 42 Motion Off Fault', class No Acknowledgement, trigger "DB302_HMI_Faults_Carrier42_Faults_2" bit 0
   2722: 'Carrier 42 Motion On Fault', class No Acknowledgement, trigger "DB302_HMI_Faults_Carrier42_Faults_2" bit 1
   2723: 'Carrier 42 Spacing Fault', class No Acknowledgement, trigger "DB302_HMI_Faults_Carrier42_Faults_2" bit 2
   2724: 'Carrier 42 Duplicate Carrier Number Fault', class No Acknowledgement, trigger "DB302_HMI_Faults_Carrier42_Faults_2" bit 3
   2725: 'Spare_Fault_2725', class No Acknowledgement, trigger "DB302_HMI_Faults_Carrier42_Faults_2" bit 4
   2726: 'Spare_Fault_2726', class No Acknowledgement, trigger "DB302_HMI_Faults_Carrier42_Faults_2" bit 5
   2727: 'Spare_Fault_2727', class No Acknowledgement, trigger "DB302_HMI_Faults_Carrier42_Faults_2" bit 6
   2728: 'Spare_Fault_2728', class No Acknowledgement, trigger "DB302_HMI_Faults_Carrier42_Faults_2" bit 7
   2729: 'Spare_Fault_2729', class No Acknowledgement, trigger "DB302_HMI_Faults_Carrier42_Faults_2" bit 8
   2730: 'Spare_Fault_2730', class No Acknowledgement, trigger "DB302_HMI_Faults_Carrier42_Faults_2" bit 9
   2731: 'Spare_Fault_2731', class No Acknowledgement, trigger "DB302_HMI_Faults_Carrier42_Faults_2" bit 10
   2732: 'Spare_Fault_2732', class No Acknowledgement, trigger "DB302_HMI_Faults_Carrier42_Faults_2" bit 11
   2733: 'Spare_Fault_2733', class No Acknowledgement, trigger "DB302_HMI_Faults_Carrier42_Faults_2" bit 12
   2734: 'Spare_Fault_2734', class No Acknowledgement, trigger "DB302_HMI_Faults_Carrier42_Faults_2" bit 13
   2735: 'Spare_Fault_2735', class No Acknowledgement, trigger "DB302_HMI_Faults_Carrier42_Faults_2" bit 14
   2736: 'Spare_Fault_2736', class No Acknowledgement, trigger "DB302_HMI_Faults_Carrier42_Faults_2" bit 15
   2737: 'Spare_Fault_2737', class No Acknowledgement, trigger "DB302_HMI_Faults_Carrier42_Faults_3" bit 0
   2738: 'Spare_Fault_2738', class No Acknowledgement, trigger "DB302_HMI_Faults_Carrier42_Faults_3" bit 1
   2739: 'Spare_Fault_2739', class No Acknowledgement, trigger "DB302_HMI_Faults_Carrier42_Faults_3" bit 2
   2740: 'Spare_Fault_2740', class No Acknowledgement, trigger "DB302_HMI_Faults_Carrier42_Faults_3" bit 3
   2741: 'Spare_Fault_2741', class No Acknowledgement, trigger "DB302_HMI_Faults_Carrier42_Faults_3" bit 4
   2742: 'Spare_Fault_2742', class No Acknowledgement, trigger "DB302_HMI_Faults_Carrier42_Faults_3" bit 5
   2743: 'Spare_Fault_2743', class No Acknowledgement, trigger "DB302_HMI_Faults_Carrier42_Faults_3" bit 6
   2744: 'Spare_Fault_2744', class No Acknowledgement, trigger "DB302_HMI_Faults_Carrier42_Faults_3" bit 7
   2745: 'Spare_Fault_2745', class No Acknowledgement, trigger "DB302_HMI_Faults_Carrier42_Faults_3" bit 8
   2746: 'Spare_Fault_2746', class No Acknowledgement, trigger "DB302_HMI_Faults_Carrier42_Faults_3" bit 9
   2747: 'Spare_Fault_2747', class No Acknowledgement, trigger "DB302_HMI_Faults_Carrier42_Faults_3" bit 10
   2748: 'Spare_Fault_2748', class No Acknowledgement, trigger "DB302_HMI_Faults_Carrier42_Faults_3" bit 11
   2749: 'Spare_Fault_2749', class No Acknowledgement, trigger "DB302_HMI_Faults_Carrier42_Faults_3" bit 12
   2750: 'Spare_Fault_2750', class No Acknowledgement, trigger "DB302_HMI_Faults_Carrier42_Faults_3" bit 13
   2751: 'Spare_Fault_2751', class No Acknowledgement, trigger "DB302_HMI_Faults_Carrier42_Faults_3" bit 14
   2752: 'Spare_Fault_2752', class No Acknowledgement, trigger "DB302_HMI_Faults_Carrier42_Faults_3" bit 15
   2753: 'Carrier 43 Disconnect Open Power Fault DI11.0', class No Acknowledgement, trigger "DB302_HMI_Faults_Carrier43_Faults_0" bit 0
   2754: 'Carrier 43 Drive Profinet Comm Fault', class No Acknowledgement, trigger "DB302_HMI_Faults_Carrier43_Faults_0" bit 1
   2755: 'Carrier 43 Production Stop Not Reset', class No Acknowledgement, trigger "DB302_HMI_Faults_Carrier43_Faults_0" bit 2
   2756: 'Carrier 43 CB02122 Tripped', class No Acknowledgement, trigger "DB302_HMI_Faults_Carrier43_Faults_0" bit 3
   2757: 'Carrier 43 CB02123 Tripped', class No Acknowledgement, trigger "DB302_HMI_Faults_Carrier43_Faults_0" bit 4
   2758: 'Carrier 43 AUX1 CB Tripped', class No Acknowledgement, trigger "DB302_HMI_Faults_Carrier43_Faults_0" bit 5
   2759: 'Carrier 43 AUX2 CB Tripped', class No Acknowledgement, trigger "DB302_HMI_Faults_Carrier43_Faults_0" bit 6
   2760: 'Carrier 43 PLC Not Communicating', class No Acknowledgement, trigger "DB302_HMI_Faults_Carrier43_Faults_0" bit 7
   2761: 'Carrier 43 Safe Input Card Fault', class No Acknowledgement, trigger "DB302_HMI_Faults_Carrier43_Faults_0" bit 8
   2762: 'Carrier 43 Safe Output Card Fault', class No Acknowledgement, trigger "DB302_HMI_Faults_Carrier43_Faults_0" bit 9
   2763: 'Carrier 43 Standard Input Card Fault', class No Acknowledgement, trigger "DB302_HMI_Faults_Carrier43_Faults_0" bit 10
   2764: 'Carrier 43 Standard Output Card Fault', class No Acknowledgement, trigger "DB302_HMI_Faults_Carrier43_Faults_0" bit 11
   2765: 'Carrier 43 Encoder Position Fault', class No Acknowledgement, trigger "DB302_HMI_Faults_Carrier43_Faults_0" bit 12
   2766: 'Carrier 43 Encoder Internal Error', class No Acknowledgement, trigger "DB302_HMI_Faults_Carrier43_Faults_0" bit 13
   2767: 'Carrier 43 Encoder Comm Fault', class No Acknowledgement, trigger "DB302_HMI_Faults_Carrier43_Faults_0" bit 14
   2768: 'Carrier 43 HMI Comm Fault', class No Acknowledgement, trigger "DB302_HMI_Faults_Carrier43_Faults_0" bit 15
   2769: 'Carrier 43 Crash Detection Fault', class No Acknowledgement, trigger "DB302_HMI_Faults_Carrier43_Faults_1" bit 0
   2770: 'Carrier 43 Carrier Number Invalid', class No Acknowledgement, trigger "DB302_HMI_Faults_Carrier43_Faults_1" bit 1
   2771: 'Carrier 43 Drive: PROFINET configuration error', class No Acknowledgement, trigger "DB302_HMI_Faults_Carrier43_Faults_1" bit 2
   2772: 'Carrier 43 Drive: Error internal communications', class No Acknowledgement, trigger "DB302_HMI_Faults_Carrier43_Faults_1" bit 3
   2773: 'Carrier 43 Drive: Motor overtemperature', class No Acknowledgement, trigger "DB302_HMI_Faults_Carrier43_Faults_1" bit 4
   2774: 'Carrier 43 Drive: Motor overcurrent', class No Acknowledgement, trigger "DB302_HMI_Faults_Carrier43_Faults_1" bit 5
   2775: 'Carrier 43 Drive: Infeed or power unit not ready', class No Acknowledgement, trigger "DB302_HMI_Faults_Carrier43_Faults_1" bit 6
   2776: 'Carrier 43 Drive: Short-circuit/ground fault detected', class No Acknowledgement, trigger "DB302_HMI_Faults_Carrier43_Faults_1" bit 7
   2777: 'Carrier 43 Drive: PROFINET Setpoint timeout', class No Acknowledgement, trigger "DB302_HMI_Faults_Carrier43_Faults_1" bit 8
   2778: 'Carrier 43 Power unit: Overcurrent', class No Acknowledgement, trigger "DB302_HMI_Faults_Carrier43_Faults_1" bit 9
   2779: 'Carrier 43 Power unit: DC link voltage overvoltage', class No Acknowledgement, trigger "DB302_HMI_Faults_Carrier43_Faults_1" bit 10
   2780: 'Carrier 43 Power unit: DC link voltage undervoltage', class No Acknowledgement, trigger "DB302_HMI_Faults_Carrier43_Faults_1" bit 11
   2781: 'Carrier 43 Power unit: Line phase failure in main circuit', class No Acknowledgement, trigger "DB302_HMI_Faults_Carrier43_Faults_1" bit 12
   2782: 'Carrier 43 Power unit: Phase failure motor cable', class No Acknowledgement, trigger "DB302_HMI_Faults_Carrier43_Faults_1" bit 13
   2783: 'Carrier 43 Power unit: Ground fault', class No Acknowledgement, trigger "DB302_HMI_Faults_Carrier43_Faults_1" bit 14
   2784: 'Spare_Fault_2784', class No Acknowledgement, trigger "DB302_HMI_Faults_Carrier43_Faults_1" bit 15
   2785: 'Carrier 43 Motion Off Fault', class No Acknowledgement, trigger "DB302_HMI_Faults_Carrier43_Faults_2" bit 0
   2786: 'Carrier 43 Motion On Fault', class No Acknowledgement, trigger "DB302_HMI_Faults_Carrier43_Faults_2" bit 1
   2787: 'Carrier 43 Spacing Fault', class No Acknowledgement, trigger "DB302_HMI_Faults_Carrier43_Faults_2" bit 2
   2788: 'Carrier 43 Duplicate Carrier Number Fault', class No Acknowledgement, trigger "DB302_HMI_Faults_Carrier43_Faults_2" bit 3
   2789: 'Spare_Fault_2789', class No Acknowledgement, trigger "DB302_HMI_Faults_Carrier43_Faults_2" bit 4
   2790: 'Spare_Fault_2790', class No Acknowledgement, trigger "DB302_HMI_Faults_Carrier43_Faults_2" bit 5
   2791: 'Spare_Fault_2791', class No Acknowledgement, trigger "DB302_HMI_Faults_Carrier43_Faults_2" bit 6
   2792: 'Spare_Fault_2792', class No Acknowledgement, trigger "DB302_HMI_Faults_Carrier43_Faults_2" bit 7
   2793: 'Spare_Fault_2793', class No Acknowledgement, trigger "DB302_HMI_Faults_Carrier43_Faults_2" bit 8
   2794: 'Spare_Fault_2794', class No Acknowledgement, trigger "DB302_HMI_Faults_Carrier43_Faults_2" bit 9
   2795: 'Spare_Fault_2795', class No Acknowledgement, trigger "DB302_HMI_Faults_Carrier43_Faults_2" bit 10
   2796: 'Spare_Fault_2796', class No Acknowledgement, trigger "DB302_HMI_Faults_Carrier43_Faults_2" bit 11
   2797: 'Spare_Fault_2797', class No Acknowledgement, trigger "DB302_HMI_Faults_Carrier43_Faults_2" bit 12
   2798: 'Spare_Fault_2798', class No Acknowledgement, trigger "DB302_HMI_Faults_Carrier43_Faults_2" bit 13
   2799: 'Spare_Fault_2799', class No Acknowledgement, trigger "DB302_HMI_Faults_Carrier43_Faults_2" bit 14
   2800: 'Spare_Fault_2800', class No Acknowledgement, trigger "DB302_HMI_Faults_Carrier43_Faults_2" bit 15
   2801: 'Spare_Fault_2801', class No Acknowledgement, trigger "DB302_HMI_Faults_Carrier43_Faults_3" bit 0
   2802: 'Spare_Fault_2802', class No Acknowledgement, trigger "DB302_HMI_Faults_Carrier43_Faults_3" bit 1
   2803: 'Spare_Fault_2803', class No Acknowledgement, trigger "DB302_HMI_Faults_Carrier43_Faults_3" bit 2